(* Logix 5000 project; controller FV vendor 1 type 14 code 217 rev 31.11; software revision 31.00; part 59 of 63 *)
(* tags used below, declared in another part *)
   Alarm_Reset : BOOL;
   Analog_Fault_No : DINT;
   Analog_Simulation_Enabled : BOOL;
   CWD : CHECKWORD_FLAGS;
   Default_Check_Time : DINT;
   FtoF_raw_input : REAL;
   Item_Simulation_Flag : BOOL;
   ItoF_raw_input : INT;
   One_Second_One_Scan : ALIAS FOR One_Second_1_scan;
   overrange_RIO_analog_value : REAL;
   rack_simulation_flag : BOOL;
   Scada_Pump_Fault_No : DINT;
   Scada_Pump_H_Fault_No : DINT;
   Scada_Pump_T_Fault_No : DINT;
   Scada_Valve_Fault_No : DINT;
   scale_analog_int : DINT;
   scale_analog_result : REAL;
   scale_eu_max : REAL;
   scale_eu_min : REAL;
   scale_raw_input : REAL;
   scale_raw_max : REAL;
   scale_raw_min : REAL;
   scale_routine_active : BOOL;
   scale_temp : REAL;
   template_analog_input : PlantItem;
   template_analog_input_RawInput : REAL;
   template_analog_output : PlantItem;
   template_analog_output_RawOutput : REAL;
   template_input : PlantItem;
   template_input_RawInput : ALIAS FOR template_boolean;
   template_output : PlantItem;
   template_output_RawOutput : ALIAS FOR template_boolean;   // P04CHILLRUN Chiller Run Signal
   template_pump : PlantItem;
   template_pump_D : ALIAS FOR template_boolean;   // auto start vacuum pump 1
   template_pump_ISOL : ALIAS FOR template_boolean;
   template_pump_R : ALIAS FOR template_boolean;   // vacuum pump 1 running
   template_valve : PlantItem;
   template_valve_C : ALIAS FOR template_boolean;   // skim manifold to ycv2 drain valve closed
   template_valve_DR : ALIAS FOR template_boolean;   // drive open skim manifold to ycv2 drain valve
   template_valve_O : ALIAS FOR template_boolean;   // skim manifold to ycv2 drain valve opened
   underrange_RIO_analog_value : REAL;
   YP_B103 : INT[15];   // Original N File From SLC, No Description Available
   YP_B3 : INT[7];   // BINARY
   YP_B30 : INT[37];   // Original N File From SLC, No Description Available
   YP_B92 : INT[105];   // Original N File From SLC, No Description Available
   YP_N7 : INT[56];   // INTEGER
   YP_T20 : TIMER[55];

PROGRAM Last_Task   (* main routine MainRoutine *)

ROUTINE MainRoutine   (* ladder *)
   0: NOP();
END_ROUTINE
END_PROGRAM

PROGRAM Templates   (* main routine Normal_Input_Template *)

ROUTINE Analog_Scale_FtoI   (* ladder *)
   0: SBR(scale_raw_input,scale_raw_min,scale_raw_max,scale_eu_min,scale_eu_max)OTE(scale_routine_active);
   1: CPT(scale_temp,(scale_eu_max-scale_eu_min)/(scale_raw_max-scale_raw_min));
   2: CPT(scale_analog_result,(scale_raw_input-scale_raw_min)*scale_temp+scale_eu_min);
   3: ADD(scale_analog_result,0.0,scale_analog_int);
   4: RET(scale_analog_int);
END_ROUTINE

ROUTINE Analog_Scale_ItoF   (* ladder *)
   0: SBR(ItoF_raw_input,scale_raw_min,scale_raw_max,scale_eu_min,scale_eu_max)OTE(scale_routine_active);
   1: ADD(ItoF_raw_input,0.0,scale_raw_input);
   2: CPT(scale_temp,(scale_eu_max-scale_eu_min)/(scale_raw_max-scale_raw_min));
   3: CPT(scale_analog_result,(scale_raw_input-scale_raw_min)*scale_temp+scale_eu_min);
   4: RET(scale_analog_result);
END_ROUTINE

ROUTINE Normal_Analogue_Input   (* ladder *)
   0: XIO(Analog_Simulation_Enabled)[XIO(template_analog_input.CW.[CWD.MANUAL]) JSR(Analog_Scale_ItoF,5,template_analog_input_RawInput,0.0,30840.0,0.0,6500.0,template_analog_input.Scaled) ,[LIM(underrange_RIO_analog_value,template_analog_input_RawInput,overrange_RIO_analog_value) ,XIC(template_analog_input.CW.[CWD.CHECKOFF]) ] CLR(template_analog_input.CheckTimer) ,XIC(S:FS) [OTU(template_analog_input.CW.[CWD.MANUAL]) ,LEQ(template_analog_input.CheckTime,0) MOV(Default_Check_Time,template_analog_input.CheckTime) ] ,XIC(One_Second_One_Scan) LES(template_analog_input.CheckTimer,template_analog_input.CheckTime) ADD(template_analog_input.CheckTimer,1,template_analog_input.CheckTimer) ,GEQ(template_analog_input.CheckTimer,template_analog_input.CheckTime) XIO(Alarm_Reset) OTE(template_analog_input.CW.[CWD.FAULT]) ,XIC(template_analog_input.CW.[CWD.FAULT]) EQU(Analog_Fault_No,0) XIO(template_analog_input.CW.[CWD.FAULTLOGGED]) [MOV(30001,Analog_Fault_No) ,OTL(template_analog_input.CW.[CWD.FAULTLOGGED]) ] ];
END_ROUTINE

ROUTINE Normal_Analogue_Output   (* ladder *)
   0: XIO(Analog_Simulation_Enabled)JSR(Analog_Scale_FtoI,5,template_analog_output.Scaled,0.0,100.0,0.0,30840.0,template_analog_output_RawOutput);
END_ROUTINE

ROUTINE Normal_Input_Template   (* ladder *)
   0: [XIC(S:FS) OTU(template_input.CW.[CWD.MANUAL]) ,[XIC(template_input_RawInput) XIO(template_input.CW.[CWD.MANUAL]) ,XIC(template_input.CW.[CWD.MANDRV]) XIC(template_input.CW.[CWD.MANUAL]) ] OTE(template_input.CW.[CWD.INPUTSTATUS]) ,XIC(One_Second_One_Scan) [XIC(template_input.CW.[CWD.INPUTSTATUS]) XIO(template_input.CW.[CWD.INPUTSTATUSDEBOUNCED]) ,XIO(template_input.CW.[CWD.INPUTSTATUS]) XIC(template_input.CW.[CWD.INPUTSTATUSDEBOUNCED]) ] ADD(1,template_input.DebounceTimer,template_input.DebounceTimer) ,[XIC(template_input.CW.[CWD.INPUTSTATUS]) XIC(template_input.CW.[CWD.INPUTSTATUSDEBOUNCED]) ,XIO(template_input.CW.[CWD.INPUTSTATUS]) XIO(template_input.CW.[CWD.INPUTSTATUSDEBOUNCED]) ] CLR(template_input.DebounceTimer) ,GEQ(template_input.DebounceTimer,template_input.DebounceTime) XIC(template_input.CW.[CWD.INPUTSTATUS]) [OTL(template_input.CW.[CWD.INPUTSTATUSDEBOUNCED]) ,CLR(template_input.DebounceTimer) ] ,GEQ(template_input.DebounceTimer,template_input.DebounceTime) XIO(template_input.CW.[CWD.INPUTSTATUS]) [OTU(template_input.CW.[CWD.INPUTSTATUSDEBOUNCED]) ,CLR(template_input.DebounceTimer) ] ];
END_ROUTINE

ROUTINE Normal_Output_Template   (* ladder *)
   0: [NEQ(template_output.DriveBits,0) OTE(template_output.CW.[CWD.AUTODRV]) ,XIC(S:FS) OTU(template_output.CW.[CWD.MANUAL]) ,[XIC(template_output.CW.[CWD.AUTODRV]) XIO(template_output.CW.[CWD.MANUAL]) ,XIC(template_output.CW.[CWD.MANDRV]) XIC(template_output.CW.[CWD.MANUAL]) ] OTE(template_output.CW.[CWD.OUTPUT]) ,XIC(template_output.CW.[CWD.OUTPUT]) OTE(template_output_RawOutput) ];
END_ROUTINE

ROUTINE Normal_Pump_Template_Isol   (* ladder *)
   0: [NEQ(template_pump.DriveBits,0) OTE(template_pump.CW.[CWD.AUTODRV]) ,[XIC(template_pump.CW.[CWD.AUTODRV]) XIO(template_pump.CW.[CWD.MANUAL]) ,XIC(template_pump.CW.[CWD.MANDRV]) XIC(template_pump.CW.[CWD.MANUAL]) ] OTE(template_pump.CW.[CWD.OUTPUT]) ,XIC(template_pump.CW.[CWD.OUTPUT]) OTE(template_pump_D) ,XIC(S:FS) [OTU(template_pump.CW.[CWD.MANUAL]) ,LEQ(template_pump.CheckTime,0) MOV(Default_Check_Time,template_pump.CheckTime) ] ,[[XIC(template_pump_R) XIO(Item_Simulation_Flag) ,XIC(Item_Simulation_Flag) [XIC(template_pump.CW.[CWD.AUTODRV]) XIO(template_pump.CW.[CWD.SIMFAIL]) ,XIO(template_pump.CW.[CWD.AUTODRV]) XIC(template_pump.CW.[CWD.SIMFAIL]) ] ] OTE(template_pump.CW.[CWD.RUNFB]) ,[XIC(rack_simulation_flag) ,XIC(template_pump.CW.[CWD.CHECKOFF]) ,XIC(template_pump_ISOL) ] OTE(template_pump.CW.[CWD.HEALTHYFB]) ] ,[XIC(template_pump.CW.[CWD.AUTODRV]) XIO(template_pump.CW.[CWD.PREVSCAN]) ,XIO(template_pump.CW.[CWD.AUTODRV]) XIC(template_pump.CW.[CWD.PREVSCAN]) ] CLR(template_pump.CheckTimer) ,XIC(One_Second_One_Scan) LES(template_pump.CheckTimer,template_pump.CheckTime) ADD(template_pump.CheckTimer,1,template_pump.CheckTimer) ,XIO(template_pump.CW.[CWD.FAULT]) OTU(template_pump.CW.[CWD.FAULTLOGGED]) ,[GEQ(template_pump.CheckTimer,template_pump.CheckTime) [XIC(template_pump.CW.[CWD.OUTPUT]) XIO(template_pump.CW.[CWD.RUNFB]) ,XIO(template_pump.CW.[CWD.OUTPUT]) XIC(template_pump.CW.[CWD.RUNFB]) ] ,XIO(template_pump.CW.[CWD.HEALTHYFB]) ,XIC(template_pump.CW.[CWD.FAULT]) ,XIC(template_pump.CW.[CWD.HIGHLIGHT]) ] XIO(template_pump.CW.[CWD.CHECKOFF]) XIO(Alarm_Reset) OTE(template_pump.CW.[CWD.FAULT]) ,XIC(template_pump.CW.[CWD.OUTPUT]) OTE(template_pump.CW.[CWD.PREVSCAN]) ,XIC(template_pump.CW.[CWD.FAULT]) EQU(Scada_Pump_Fault_No,0) XIO(template_pump.CW.[CWD.FAULTLOGGED]) [MOV(20001,Scada_Pump_Fault_No) ,OTL(template_pump.CW.[CWD.FAULTLOGGED]) ] ,XIO(template_pump.CW.[CWD.HEALTHYFB]) EQU(Scada_Pump_H_Fault_No,0) XIO(template_pump.CW.[CWD.HEALTHYFAULTLOGGED]) [MOV(20001,Scada_Pump_H_Fault_No) ,OTL(template_pump.CW.[CWD.HEALTHYFAULTLOGGED]) ] ,XIO(template_pump.CW.[CWD.NOTTRIPPEDFB]) EQU(Scada_Pump_H_Fault_No,0) XIO(template_pump.CW.[CWD.TRIPPEDFAULTLOGGED]) [MOV(20001,Scada_Pump_T_Fault_No) ,OTL(template_pump.CW.[CWD.TRIPPEDFAULTLOGGED]) ] ];
END_ROUTINE

ROUTINE Normal_Pump_Template_JustRun   (* ladder *)
   0: [NEQ(template_pump.DriveBits,0) OTE(template_pump.CW.[CWD.AUTODRV]) ,[XIC(template_pump.CW.[CWD.AUTODRV]) XIO(template_pump.CW.[CWD.MANUAL]) ,XIC(template_pump.CW.[CWD.MANDRV]) XIC(template_pump.CW.[CWD.MANUAL]) ] OTE(template_pump.CW.[CWD.OUTPUT]) ,XIC(template_pump.CW.[CWD.OUTPUT]) OTE(template_pump_D) ,XIC(S:FS) [OTU(template_pump.CW.[CWD.MANUAL]) ,LEQ(template_pump.CheckTime,0) MOV(Default_Check_Time,template_pump.CheckTime) ] ,[[XIC(template_pump_R) XIO(Item_Simulation_Flag) ,XIC(Item_Simulation_Flag) [XIC(template_pump.CW.[CWD.AUTODRV]) XIO(template_pump.CW.[CWD.SIMFAIL]) ,XIO(template_pump.CW.[CWD.AUTODRV]) XIC(template_pump.CW.[CWD.SIMFAIL]) ] ] OTE(template_pump.CW.[CWD.RUNFB]) ,[XIC(rack_simulation_flag) ,XIC(template_pump.CW.[CWD.CHECKOFF]) ,] OTE(template_pump.CW.[CWD.HEALTHYFB]) ] ,[XIC(template_pump.CW.[CWD.AUTODRV]) XIO(template_pump.CW.[CWD.PREVSCAN]) ,XIO(template_pump.CW.[CWD.AUTODRV]) XIC(template_pump.CW.[CWD.PREVSCAN]) ] CLR(template_pump.CheckTimer) ,XIC(One_Second_One_Scan) LES(template_pump.CheckTimer,template_pump.CheckTime) ADD(template_pump.CheckTimer,1,template_pump.CheckTimer) ,XIO(template_pump.CW.[CWD.FAULT]) OTU(template_pump.CW.[CWD.FAULTLOGGED]) ,[GEQ(template_pump.CheckTimer,template_pump.CheckTime) [XIC(template_pump.CW.[CWD.OUTPUT]) XIO(template_pump.CW.[CWD.RUNFB]) ,XIO(template_pump.CW.[CWD.OUTPUT]) XIC(template_pump.CW.[CWD.RUNFB]) ] ,XIO(template_pump.CW.[CWD.HEALTHYFB]) ,XIC(template_pump.CW.[CWD.FAULT]) ,XIC(template_pump.CW.[CWD.HIGHLIGHT]) ] XIO(template_pump.CW.[CWD.CHECKOFF]) XIO(Alarm_Reset) OTE(template_pump.CW.[CWD.FAULT]) ,XIC(template_pump.CW.[CWD.OUTPUT]) OTE(template_pump.CW.[CWD.PREVSCAN]) ,XIC(template_pump.CW.[CWD.FAULT]) EQU(Scada_Pump_Fault_No,0) XIO(template_pump.CW.[CWD.FAULTLOGGED]) [MOV(20001,Scada_Pump_Fault_No) ,OTL(template_pump.CW.[CWD.FAULTLOGGED]) ] ,XIO(template_pump.CW.[CWD.HEALTHYFB]) EQU(Scada_Pump_H_Fault_No,0) XIO(template_pump.CW.[CWD.HEALTHYFAULTLOGGED]) [MOV(20001,Scada_Pump_H_Fault_No) ,OTL(template_pump.CW.[CWD.HEALTHYFAULTLOGGED]) ] ,XIO(template_pump.CW.[CWD.NOTTRIPPEDFB]) EQU(Scada_Pump_H_Fault_No,0) XIO(template_pump.CW.[CWD.TRIPPEDFAULTLOGGED]) [MOV(20001,Scada_Pump_T_Fault_No) ,OTL(template_pump.CW.[CWD.TRIPPEDFAULTLOGGED]) ] ];
END_ROUTINE

ROUTINE Normal_Valve_Template   (* ladder *)
   0: [NEQ(template_valve.DriveBits,0) OTE(template_valve.CW.[CWD.AUTODRV]) ,[XIC(template_valve.CW.[CWD.AUTODRV]) XIO(template_valve.CW.[CWD.MANUAL]) ,XIC(template_valve.CW.[CWD.MANDRV]) XIC(template_valve.CW.[CWD.MANUAL]) ] OTE(template_valve.CW.[CWD.OUTPUT]) ,XIC(template_valve.CW.[CWD.OUTPUT]) OTE(template_valve_DR) ,XIC(S:FS) [OTU(template_valve.CW.[CWD.MANUAL]) ,LEQ(template_valve.CheckTime,0) MOV(Default_Check_Time,template_valve.CheckTime) ] ,[[XIC(template_valve_O) XIO(Item_Simulation_Flag) ,XIC(Item_Simulation_Flag) XIC(template_valve.CW.[CWD.AUTODRV]) XIO(template_valve.CW.[CWD.SIMFAIL]) ] OTE(template_valve.CW.[CWD.OPENFB]) ,[XIC(template_valve_C) XIO(Item_Simulation_Flag) ,XIC(Item_Simulation_Flag) XIO(template_valve.CW.[CWD.AUTODRV]) XIO(template_valve.CW.[CWD.SIMFAIL]) ] OTE(template_valve.CW.[CWD.CLOSEDFB]) ] ,[XIC(template_valve.CW.[CWD.AUTODRV]) XIO(template_valve.CW.[CWD.PREVSCAN]) ,XIO(template_valve.CW.[CWD.AUTODRV]) XIC(template_valve.CW.[CWD.PREVSCAN]) ] CLR(template_valve.CheckTimer) ,XIC(One_Second_One_Scan) LES(template_valve.CheckTimer,template_valve.CheckTime) ADD(template_valve.CheckTimer,1,template_valve.CheckTimer) ,XIO(template_valve.CW.[CWD.FAULT]) OTU(template_valve.CW.[CWD.FAULTLOGGED]) ,[GEQ(template_valve.CheckTimer,template_valve.CheckTime) [XIC(template_valve.CW.[CWD.OUTPUT]) [XIO(template_valve.CW.[CWD.OPENFB]) ,XIC(template_valve.CW.[CWD.CLOSEDFB]) ] ,XIO(template_valve.CW.[CWD.OUTPUT]) [XIC(template_valve.CW.[CWD.OPENFB]) ,XIO(template_valve.CW.[CWD.CLOSEDFB]) ] ] ,XIC(template_valve.CW.[CWD.FAULT]) ,XIC(template_valve.CW.[CWD.HIGHLIGHT]) ] XIO(template_valve.CW.[CWD.CHECKOFF]) XIO(Alarm_Reset) OTE(template_valve.CW.[CWD.FAULT]) ,XIC(template_valve.CW.[CWD.OUTPUT]) OTE(template_valve.CW.[CWD.PREVSCAN]) ,XIC(template_valve.CW.[CWD.FAULT]) EQU(Scada_Valve_Fault_No,0) XIO(template_valve.CW.[CWD.FAULTLOGGED]) [MOV(10001,Scada_Valve_Fault_No) ,OTL(template_valve.CW.[CWD.FAULTLOGGED]) ] ];
END_ROUTINE
END_PROGRAM

PROGRAM YP_Common   (* main routine MainRoutine *)

ROUTINE Analog_scale_ftof   (* ladder *)
   0: SBR(FtoF_raw_input,scale_raw_min,scale_raw_max,scale_eu_min,scale_eu_max)OTE(scale_routine_active);
   1: ADD(FtoF_raw_input,0.0,scale_raw_input);
   2: CPT(scale_temp,(scale_eu_max-scale_eu_min)/(scale_raw_max-scale_raw_min));
   3: CPT(scale_analog_result,(scale_raw_input-scale_raw_min)*scale_temp+scale_eu_min);
   4: RET(scale_analog_result);
END_ROUTINE

ROUTINE Analog_Scale_FtoI   (* ladder *)
   0: SBR(scale_raw_input,scale_raw_min,scale_raw_max,scale_eu_min,scale_eu_max)OTE(scale_routine_active);
   1: CPT(scale_temp,(scale_eu_max-scale_eu_min)/(scale_raw_max-scale_raw_min));
   2: CPT(scale_analog_result,(scale_raw_input-scale_raw_min)*scale_temp+scale_eu_min);
   3: ADD(scale_analog_result,0.0,scale_analog_int);
   4: RET(scale_analog_int);
END_ROUTINE

ROUTINE Analog_Scale_ItoF   (* ladder *)
   0: SBR(ItoF_raw_input,scale_raw_min,scale_raw_max,scale_eu_min,scale_eu_max)OTE(scale_routine_active);
   1: ADD(ItoF_raw_input,0.0,scale_raw_input);
   2: CPT(scale_temp,(scale_eu_max-scale_eu_min)/(scale_raw_max-scale_raw_min));
   3: CPT(scale_analog_result,(scale_raw_input-scale_raw_min)*scale_temp+scale_eu_min);
   4: RET(scale_analog_result);
END_ROUTINE

ROUTINE Constants   (* ladder *)
   0: [MOV(0,CWD.AUTODRV) ,MOV(0,CWD.INPUTSTATUS) ,MOV(1,CWD.PREVSCAN) ,MOV(2,CWD.SIMFAIL) ,MOV(3,CWD.OPENFB) ,MOV(3,CWD.RUNFB) ,MOV(4,CWD.CLOSEDFB) ,MOV(5,CWD.MANDRV) ,MOV(6,CWD.MANUAL) ,MOV(7,CWD.OUTPUT) ,MOV(8,CWD.CHECKOFF) ,MOV(9,CWD.HIGHLIGHT) ,MOV(10,CWD.HEALTHYFB) ,MOV(11,CWD.NOTTRIPPEDFB) ,MOV(12,CWD.ANALOGSIMULATION) ,MOV(14,CWD.FAULTLOGGED) ,MOV(15,CWD.FAULT) ,MOV(16,CWD.HEALTHYFAULTLOGGED) ,MOV(17,CWD.TRIPPEDFAULTLOGGED) ];
END_ROUTINE

ROUTINE MainRoutine   (* ladder *)
   0: XIC(s:fs)JSR(Constants,0);
   // Always Force Alarm Reset to be pushed Until Delphi Code Removed, Original Delphi did not have global alarm reset.
   1: OTU(Alarm_Reset);
   2: JSR(YP_Digital_Inputs,0);
   3: JSR(YP_Digital_Outputs,0);
   4: JSR(YP_Valves,0);
   5: JSR(YP_ALARMS_3,0);
   6: JSR(YP_COMMS_4,0);
   7: JSR(YP_INPUTS_10,0);
   8: JSR(YP_OUTPUTS_11,0);
   9: JSR(YP_BLUNGER_14,0);
   10: JSR(YP_LAD15_15,0);
   11: JSR(YP_LAD16_16,0);
   12: JSR(YP_RQD_FLAGS_17,0);
   13: JSR(YP_YSTS_HL_18,0);
   14: JSR(YP_LAD20_20,0);
END_ROUTINE

ROUTINE YP_ALARMS_3   (* ladder *)
   0: XIC(YP_B30[0].3)XIO(YP_B3[0].0)TON(YP_T20[0],?,?);
   1: XIO(YP_B30[0].3)XIC(YP_B3[0].0)TON(YP_T20[1],?,?);
   2: XIC(YP_B30[0].5)XIO(YP_B3[0].2)TON(YP_T20[2],?,?);
   3: XIO(YP_B30[0].5)XIC(YP_B3[0].2)TON(YP_T20[3],?,?);
   4: XIC(YP_B30[0].6)XIO(YP_B3[0].4)TON(YP_T20[4],?,?);
   5: XIO(YP_B30[0].6)XIC(YP_B3[0].4)TON(YP_T20[5],?,?);
   6: XIC(YP_B30[0].7)XIO(YP_B3[0].6)TON(YP_T20[6],?,?);
   7: XIO(YP_B30[0].7)XIC(YP_B3[0].6)TON(YP_T20[7],?,?);
   8: XIC(YP_B30[0].8)XIO(YP_B3[0].8)TON(YP_T20[8],?,?);
   9: XIO(YP_B30[0].8)XIC(YP_B3[0].8)TON(YP_T20[9],?,?);
   10: XIC(YP_B30[0].9)XIO(YP_B3[0].10)TON(YP_T20[10],?,?);
   11: XIO(YP_B30[0].9)XIC(YP_B3[0].10)TON(YP_T20[11],?,?);
   12: XIC(YP_B30[0].10)XIO(YP_B3[0].12)TON(YP_T20[12],?,?);
   13: XIO(YP_B30[0].10)XIC(YP_B3[0].12)TON(YP_T20[13],?,?);
   14: XIC(YP_B30[0].11)XIO(YP_B3[0].14)TON(YP_T20[14],?,?);
   15: XIO(YP_B30[0].11)XIC(YP_B3[0].14)TON(YP_T20[15],?,?);
   16: XIC(YP_B30[0].1)TON(YP_T20[16],?,?);
   17: XIC(YP_B30[0].0)TON(YP_T20[17],?,?);
   18: XIC(YP_B103[0].0)TON(YP_T20[18],?,?);
   19: XIC(YP_T20[0].DN)OTE(YP_B92[0].0);
   20: XIC(YP_T20[1].DN)OTE(YP_B92[0].1);
   21: XIC(YP_T20[2].DN)OTE(YP_B92[0].2);
   22: XIC(YP_T20[3].DN)OTE(YP_B92[0].3);
   23: XIC(YP_T20[4].DN)OTE(YP_B92[0].4);
   24: XIC(YP_T20[5].DN)OTE(YP_B92[0].5);
   25: XIC(YP_T20[6].DN)OTE(YP_B92[0].6);
   26: XIC(YP_T20[7].DN)OTE(YP_B92[0].7);
   27: XIC(YP_T20[8].DN)OTE(YP_B92[0].8);
   28: XIC(YP_T20[9].DN)OTE(YP_B92[0].9);
   29: XIC(YP_T20[10].DN)OTE(YP_B92[0].10);
   30: XIC(YP_T20[11].DN)OTE(YP_B92[0].11);
   31: XIC(YP_T20[12].DN)OTE(YP_B92[0].12);
   32: XIC(YP_T20[13].DN)OTE(YP_B92[0].13);
   33: XIC(YP_T20[14].DN)OTE(YP_B92[0].14);
   34: XIC(YP_T20[15].DN)OTE(YP_B92[0].15);
   35: XIC(YP_N7[38].0)OTE(YP_B92[1].0);
   36: XIC(YP_N7[38].1)OTE(YP_B92[1].1);
   37: XIC(YP_B3[1].13)OTE(YP_B92[1].7);
   38: XIC(YP_B3[1].8)OTE(YP_B92[1].10);
   39: XIC(YP_B3[1].9)OTE(YP_B92[1].11);
   40: XIC(YP_T20[16].DN)OTE(YP_B92[2].0);
   41: XIC(YP_T20[17].DN)OTE(YP_B92[2].1);
   42: XIC(YP_T20[18].DN)OTE(YP_B92[2].2);
   43: [AND(YP_B92[0],YP_B92[40],YP_B92[40]) ,OR(YP_B92[0],YP_B92[20],YP_B92[60]) ,XOR(YP_B92[40],YP_B92[60],YP_B92[20]) ];
   44: [AND(YP_B92[1],YP_B92[41],YP_B92[41]) ,OR(YP_B92[1],YP_B92[21],YP_B92[61]) ,XOR(YP_B92[41],YP_B92[61],YP_B92[21]) ];
   45: [AND(YP_B92[2],YP_B92[42],YP_B92[42]) ,OR(YP_B92[2],YP_B92[22],YP_B92[62]) ,XOR(YP_B92[42],YP_B92[62],YP_B92[22]) ];
   46: [AND(YP_B92[3],YP_B92[43],YP_B92[43]) ,OR(YP_B92[3],YP_B92[23],YP_B92[63]) ,XOR(YP_B92[43],YP_B92[63],YP_B92[23]) ];
